REGION Network 8: END: Update the ENO Output. (DO NOT REMOVE. Must be last rung)
   RUNG wire#powerrail
      ReturnCoil( TRUE )
   END_RUNG
   // the same network as SCL:
   ENO := TRUE;
   RETURN;
END_REGION
END_FUNCTION_BLOCK

FUNCTION_BLOCK "UN_07_RecipeControl"   // FB31627, LAD
TITLE = UN_07_RecipeControl
{ S7_Optimized_Access := 'TRUE' }
AUTHOR : tech.team.motioncontrol@siemens.com
FAMILY : CPG
VERSION : 1.0
// Support: tech.team.motioncontrol@siemens.com
   VAR
      instRecipeControl : "CPG_RecipeControl";
      instRecipeManager : "CPG_RecipeHMIManager";
      ONS_RecipeChange : Bool;
      ONS_SaveAsChange : Bool;
      ONS_DeleteChange : Bool;
      ONS_CopyChange : Bool;
   END_VAR
   VAR_TEMP
      tempEnablechange : Bool;
      tempRecipenewname : String[60];
      tempErrorID : Word;
      tempError : Word;
      tempSeconds : Time;
   END_VAR
   VAR CONSTANT
      ERR_CHANGE : Word := 16#8001;
      ERR_SAVE : Word := 16#8002;
      ERR_COPY : Word := 16#8004;
      ERR_DELETE : Word := 16#8008;
   END_VAR
   VAR_TEMP   // added for the SCL form of the ladder/FBD networks
      _w1 : Bool;
      _w2 : Bool;
   END_VAR
BEGIN

REGION Network 1: Determine if recipe change is permitted based on machine state
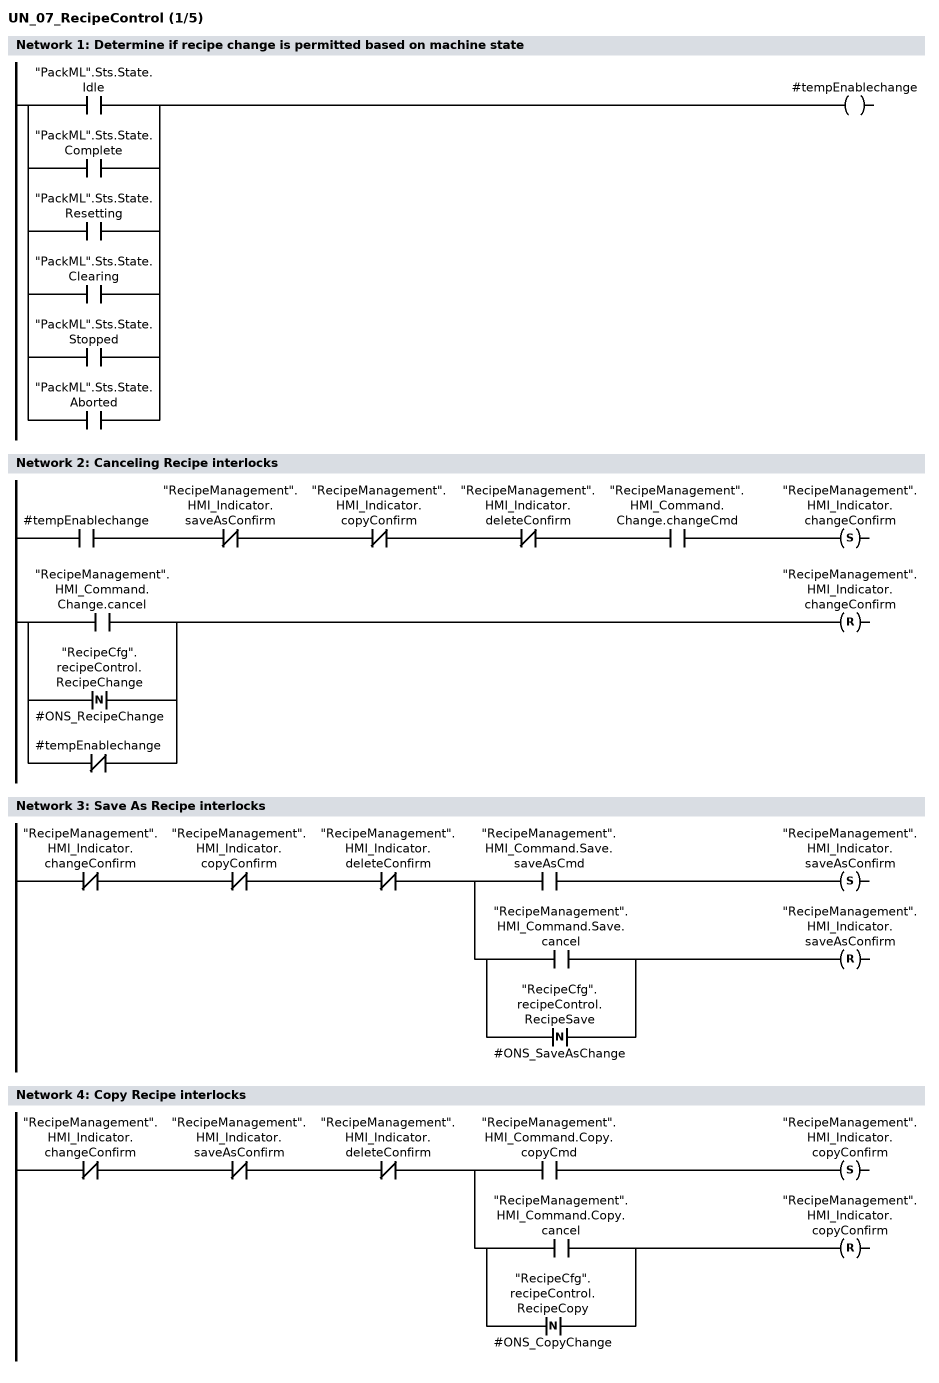
   RUNG wire#powerrail
      Contact( "PackML".Sts.State.Idle )
      wire#w1
      Coil( #tempEnablechange )
   END_RUNG
   RUNG wire#powerrail
      Contact( "PackML".Sts.State.Complete )
   END_RUNG wire#w1
   RUNG wire#powerrail
      Contact( "PackML".Sts.State.Resetting )
   END_RUNG wire#w1
   RUNG wire#powerrail
      Contact( "PackML".Sts.State.Clearing )
   END_RUNG wire#w1
   RUNG wire#powerrail
      Contact( "PackML".Sts.State.Stopped )
   END_RUNG wire#w1
   RUNG wire#powerrail
      Contact( "PackML".Sts.State.Aborted )
   END_RUNG wire#w1
   // the same network as SCL:
   #tempEnablechange := "PackML".Sts.State.Idle OR "PackML".Sts.State.Complete OR "PackML".Sts.State.Resetting OR "PackML".Sts.State.Clearing OR "PackML".Sts.State.Stopped OR "PackML".Sts.State.Aborted;
END_REGION

REGION Network 2: Canceling Recipe interlocks
   RUNG wire#powerrail
      Contact( #tempEnablechange )
      I_Contact( "RecipeManagement".HMI_Indicator.saveAsConfirm )
      I_Contact( "RecipeManagement".HMI_Indicator.copyConfirm )
      I_Contact( "RecipeManagement".HMI_Indicator.deleteConfirm )
      Contact( "RecipeManagement".HMI_Command.Change.changeCmd )
      S_Coil( "RecipeManagement".HMI_Indicator.changeConfirm )
   END_RUNG
   RUNG wire#powerrail
      Contact( "RecipeManagement".HMI_Command.Change.cancel )
      wire#w1
      R_Coil( "RecipeManagement".HMI_Indicator.changeConfirm )
   END_RUNG
   RUNG wire#powerrail
      N_Contact(operand := "RecipeCfg".recipeControl.RecipeChange, bit := #ONS_RecipeChange)
   END_RUNG wire#w1
   RUNG wire#powerrail
      I_Contact( #tempEnablechange )
   END_RUNG wire#w1
   // the same network as SCL:
   IF #tempEnablechange AND NOT "RecipeManagement".HMI_Indicator.saveAsConfirm AND NOT "RecipeManagement".HMI_Indicator.copyConfirm AND NOT "RecipeManagement".HMI_Indicator.deleteConfirm AND "RecipeManagement".HMI_Command.Change.changeCmd THEN
       "RecipeManagement".HMI_Indicator.changeConfirm := TRUE;
   END_IF;
   #_w1 := NOT "RecipeCfg".recipeControl.RecipeChange AND #ONS_RecipeChange;   // falling edge of "RecipeCfg".recipeControl.RecipeChange
   #ONS_RecipeChange := "RecipeCfg".recipeControl.RecipeChange;
   IF "RecipeManagement".HMI_Command.Change.cancel OR #_w1 OR NOT #tempEnablechange THEN
       "RecipeManagement".HMI_Indicator.changeConfirm := FALSE;
   END_IF;
END_REGION

REGION Network 3: Save As Recipe interlocks
   RUNG wire#powerrail
      I_Contact( "RecipeManagement".HMI_Indicator.changeConfirm )
      I_Contact( "RecipeManagement".HMI_Indicator.copyConfirm )
      I_Contact( "RecipeManagement".HMI_Indicator.deleteConfirm )
      wire#w1
      Contact( "RecipeManagement".HMI_Command.Save.saveAsCmd )
      S_Coil( "RecipeManagement".HMI_Indicator.saveAsConfirm )
   END_RUNG
   RUNG wire#w1
      Contact( "RecipeManagement".HMI_Command.Save.cancel )
      wire#w2
      R_Coil( "RecipeManagement".HMI_Indicator.saveAsConfirm )
   END_RUNG
   RUNG wire#w1
      N_Contact(operand := "RecipeCfg".recipeControl.RecipeSave, bit := #ONS_SaveAsChange)
   END_RUNG wire#w2
   // the same network as SCL:
   #_w1 := NOT "RecipeManagement".HMI_Indicator.changeConfirm AND NOT "RecipeManagement".HMI_Indicator.copyConfirm AND NOT "RecipeManagement".HMI_Indicator.deleteConfirm;
   IF #_w1 AND "RecipeManagement".HMI_Command.Save.saveAsCmd THEN
       "RecipeManagement".HMI_Indicator.saveAsConfirm := TRUE;
   END_IF;
   #_w2 := #_w1 AND NOT "RecipeCfg".recipeControl.RecipeSave AND #ONS_SaveAsChange;   // falling edge of "RecipeCfg".recipeControl.RecipeSave
   #ONS_SaveAsChange := "RecipeCfg".recipeControl.RecipeSave;
   IF (#_w1 AND "RecipeManagement".HMI_Command.Save.cancel) OR #_w2 THEN
       "RecipeManagement".HMI_Indicator.saveAsConfirm := FALSE;
   END_IF;
END_REGION

REGION Network 4: Copy Recipe interlocks
   RUNG wire#powerrail
      I_Contact( "RecipeManagement".HMI_Indicator.changeConfirm )
      I_Contact( "RecipeManagement".HMI_Indicator.saveAsConfirm )
      I_Contact( "RecipeManagement".HMI_Indicator.deleteConfirm )
      wire#w1
      Contact( "RecipeManagement".HMI_Command.Copy.copyCmd )
      S_Coil( "RecipeManagement".HMI_Indicator.copyConfirm )
   END_RUNG
   RUNG wire#w1
      Contact( "RecipeManagement".HMI_Command.Copy.cancel )
      wire#w2
      R_Coil( "RecipeManagement".HMI_Indicator.copyConfirm )
   END_RUNG
   RUNG wire#w1
      N_Contact(operand := "RecipeCfg".recipeControl.RecipeCopy, bit := #ONS_CopyChange)
   END_RUNG wire#w2
   // the same network as SCL:
   #_w1 := NOT "RecipeManagement".HMI_Indicator.changeConfirm AND NOT "RecipeManagement".HMI_Indicator.saveAsConfirm AND NOT "RecipeManagement".HMI_Indicator.deleteConfirm;
   IF #_w1 AND "RecipeManagement".HMI_Command.Copy.copyCmd THEN
       "RecipeManagement".HMI_Indicator.copyConfirm := TRUE;
   END_IF;
   #_w2 := #_w1 AND NOT "RecipeCfg".recipeControl.RecipeCopy AND #ONS_CopyChange;   // falling edge of "RecipeCfg".recipeControl.RecipeCopy
   #ONS_CopyChange := "RecipeCfg".recipeControl.RecipeCopy;
   IF (#_w1 AND "RecipeManagement".HMI_Command.Copy.cancel) OR #_w2 THEN
       "RecipeManagement".HMI_Indicator.copyConfirm := FALSE;
   END_IF;
END_REGION

REGION Network 5: Delete Recipe interlocks
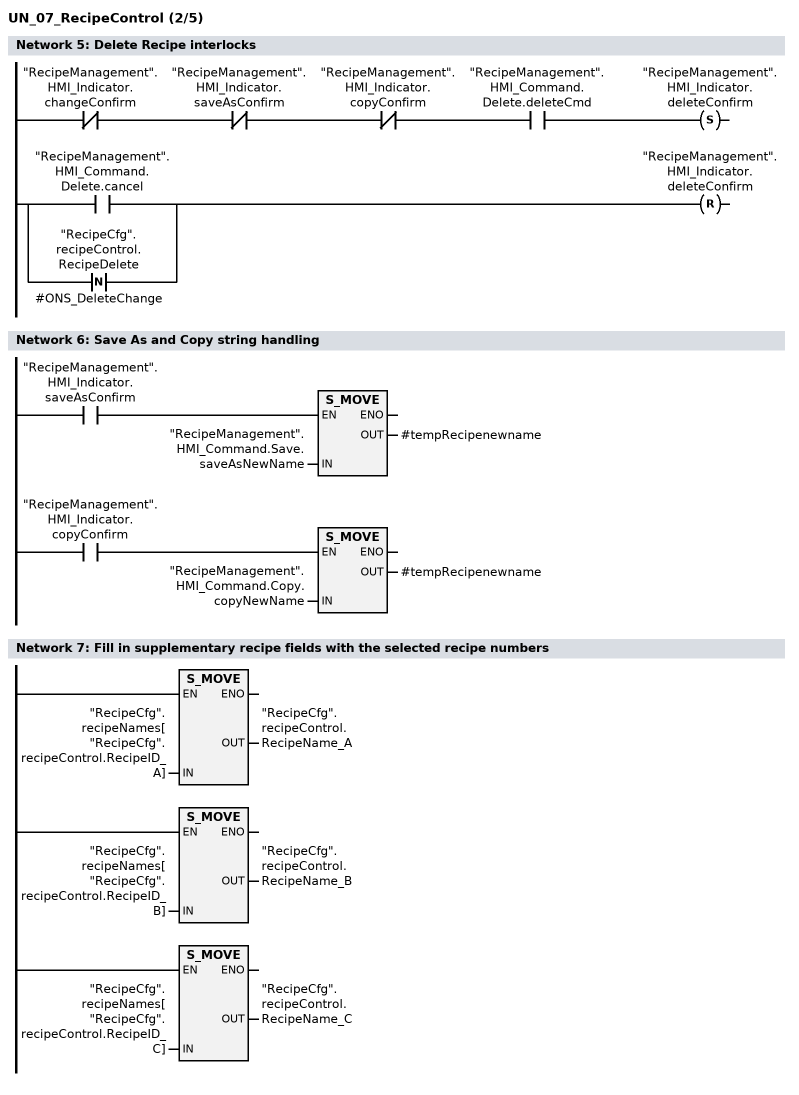
   RUNG wire#powerrail
      I_Contact( "RecipeManagement".HMI_Indicator.changeConfirm )
      I_Contact( "RecipeManagement".HMI_Indicator.saveAsConfirm )
      I_Contact( "RecipeManagement".HMI_Indicator.copyConfirm )
      Contact( "RecipeManagement".HMI_Command.Delete.deleteCmd )
      S_Coil( "RecipeManagement".HMI_Indicator.deleteConfirm )
   END_RUNG
   RUNG wire#powerrail
      Contact( "RecipeManagement".HMI_Command.Delete.cancel )
      wire#w1
      R_Coil( "RecipeManagement".HMI_Indicator.deleteConfirm )
   END_RUNG
   RUNG wire#powerrail
      N_Contact(operand := "RecipeCfg".recipeControl.RecipeDelete, bit := #ONS_DeleteChange)
   END_RUNG wire#w1
   // the same network as SCL:
   IF NOT "RecipeManagement".HMI_Indicator.changeConfirm AND NOT "RecipeManagement".HMI_Indicator.saveAsConfirm AND NOT "RecipeManagement".HMI_Indicator.copyConfirm AND "RecipeManagement".HMI_Command.Delete.deleteCmd THEN
       "RecipeManagement".HMI_Indicator.deleteConfirm := TRUE;
   END_IF;
   #_w1 := NOT "RecipeCfg".recipeControl.RecipeDelete AND #ONS_DeleteChange;   // falling edge of "RecipeCfg".recipeControl.RecipeDelete
   #ONS_DeleteChange := "RecipeCfg".recipeControl.RecipeDelete;
   IF "RecipeManagement".HMI_Command.Delete.cancel OR #_w1 THEN
       "RecipeManagement".HMI_Indicator.deleteConfirm := FALSE;
   END_IF;
END_REGION

REGION Network 6: Save As and Copy string handling
   RUNG wire#powerrail
      Contact( "RecipeManagement".HMI_Indicator.saveAsConfirm )
      S_Move(in := "RecipeManagement".HMI_Command.Save.saveAsNewName, out => #tempRecipenewname)
   END_RUNG
   RUNG wire#powerrail
      Contact( "RecipeManagement".HMI_Indicator.copyConfirm )
      S_Move(in := "RecipeManagement".HMI_Command.Copy.copyNewName, out => #tempRecipenewname)
   END_RUNG
   // the same network as SCL:
   IF "RecipeManagement".HMI_Indicator.saveAsConfirm THEN
       #tempRecipenewname := "RecipeManagement".HMI_Command.Save.saveAsNewName;
   END_IF;
   IF "RecipeManagement".HMI_Indicator.copyConfirm THEN
       #tempRecipenewname := "RecipeManagement".HMI_Command.Copy.copyNewName;
   END_IF;
END_REGION

REGION Network 7: Fill in supplementary recipe fields with the selected recipe numbers
   RUNG wire#powerrail
      S_Move(in := "RecipeCfg".recipeNames["RecipeCfg".recipeControl.RecipeID_A], out => "RecipeCfg".recipeControl.RecipeName_A)
   END_RUNG
   RUNG wire#powerrail
      S_Move(in := "RecipeCfg".recipeNames["RecipeCfg".recipeControl.RecipeID_B], out => "RecipeCfg".recipeControl.RecipeName_B)
   END_RUNG
   RUNG wire#powerrail
      S_Move(in := "RecipeCfg".recipeNames["RecipeCfg".recipeControl.RecipeID_C], out => "RecipeCfg".recipeControl.RecipeName_C)
   END_RUNG
   // the same network as SCL:
   "RecipeCfg".recipeControl.RecipeName_A := "RecipeCfg".recipeNames["RecipeCfg".recipeControl.RecipeID_A];
   "RecipeCfg".recipeControl.RecipeName_B := "RecipeCfg".recipeNames["RecipeCfg".recipeControl.RecipeID_B];
   "RecipeCfg".recipeControl.RecipeName_C := "RecipeCfg".recipeNames["RecipeCfg".recipeControl.RecipeID_C];
END_REGION

REGION Network 8: Call Recipe Control
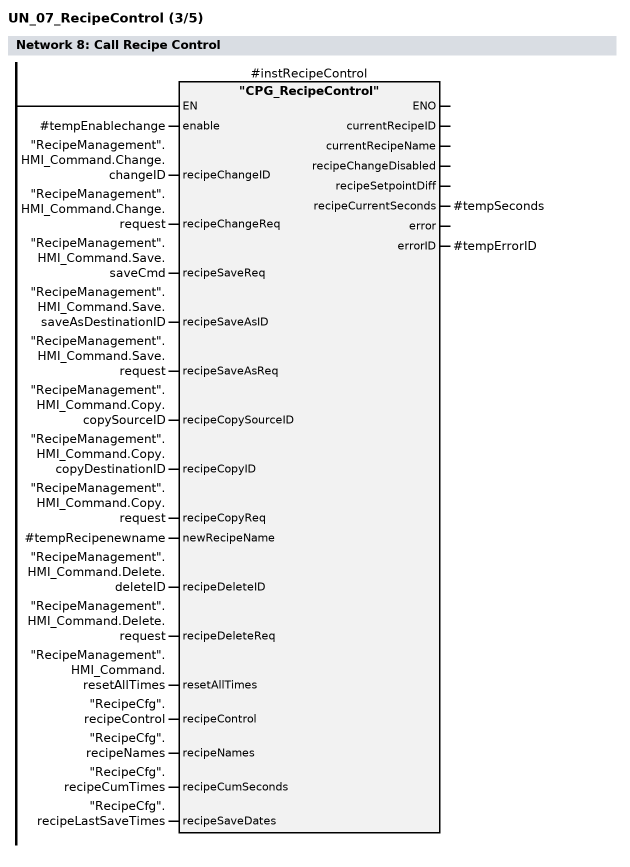
   RUNG wire#powerrail
      #instRecipeControl(enable := #tempEnablechange, recipeChangeID := "RecipeManagement".HMI_Command.Change.changeID, recipeChangeReq := "RecipeManagement".HMI_Command.Change.request, recipeSaveReq := "RecipeManagement".HMI_Command.Save.saveCmd, recipeSaveAsID := "RecipeManagement".HMI_Command.Save.saveAsDestinationID, recipeSaveAsReq := "RecipeManagement".HMI_Command.Save.request, recipeCopySourceID := "RecipeManagement".HMI_Command.Copy.copySourceID, recipeCopyID := "RecipeManagement".HMI_Command.Copy.copyDestinationID, recipeCopyReq := "RecipeManagement".HMI_Command.Copy.request, newRecipeName := #tempRecipenewname, recipeDeleteID := "RecipeManagement".HMI_Command.Delete.deleteID, recipeDeleteReq := "RecipeManagement".HMI_Command.Delete.request, resetAllTimes := "RecipeManagement".HMI_Command.resetAllTimes, recipeControl := "RecipeCfg".recipeControl, recipeNames := "RecipeCfg".recipeNames, recipeCumSeconds := "RecipeCfg".recipeCumTimes, recipeSaveDates := "RecipeCfg".recipeLastSaveTimes, currentRecipeID =>, currentRecipeName =>, recipeChangeDisabled =>, recipeSetpointDiff =>, recipeCurrentSeconds => #tempSeconds, error =>, errorID => #tempErrorID)
   END_RUNG
   // the same network as SCL:
   #instRecipeControl(enable := #tempEnablechange,   // "CPG_RecipeControl"
                      recipeChangeID := "RecipeManagement".HMI_Command.Change.changeID,
                      recipeChangeReq := "RecipeManagement".HMI_Command.Change.request,
                      recipeSaveReq := "RecipeManagement".HMI_Command.Save.saveCmd,
                      recipeSaveAsID := "RecipeManagement".HMI_Command.Save.saveAsDestinationID,
                      recipeSaveAsReq := "RecipeManagement".HMI_Command.Save.request,
                      recipeCopySourceID := "RecipeManagement".HMI_Command.Copy.copySourceID,
                      recipeCopyID := "RecipeManagement".HMI_Command.Copy.copyDestinationID,
                      recipeCopyReq := "RecipeManagement".HMI_Command.Copy.request,
                      newRecipeName := #tempRecipenewname,
                      recipeDeleteID := "RecipeManagement".HMI_Command.Delete.deleteID,
                      recipeDeleteReq := "RecipeManagement".HMI_Command.Delete.request,
                      resetAllTimes := "RecipeManagement".HMI_Command.resetAllTimes,
                      recipeControl := "RecipeCfg".recipeControl,
                      recipeNames := "RecipeCfg".recipeNames,
                      recipeCumSeconds := "RecipeCfg".recipeCumTimes,
                      recipeSaveDates := "RecipeCfg".recipeLastSaveTimes,
                      recipeCurrentSeconds => #tempSeconds,
                      errorID => #tempErrorID);
END_REGION

REGION Network 9: Clear IDs from HMI if not on that screen
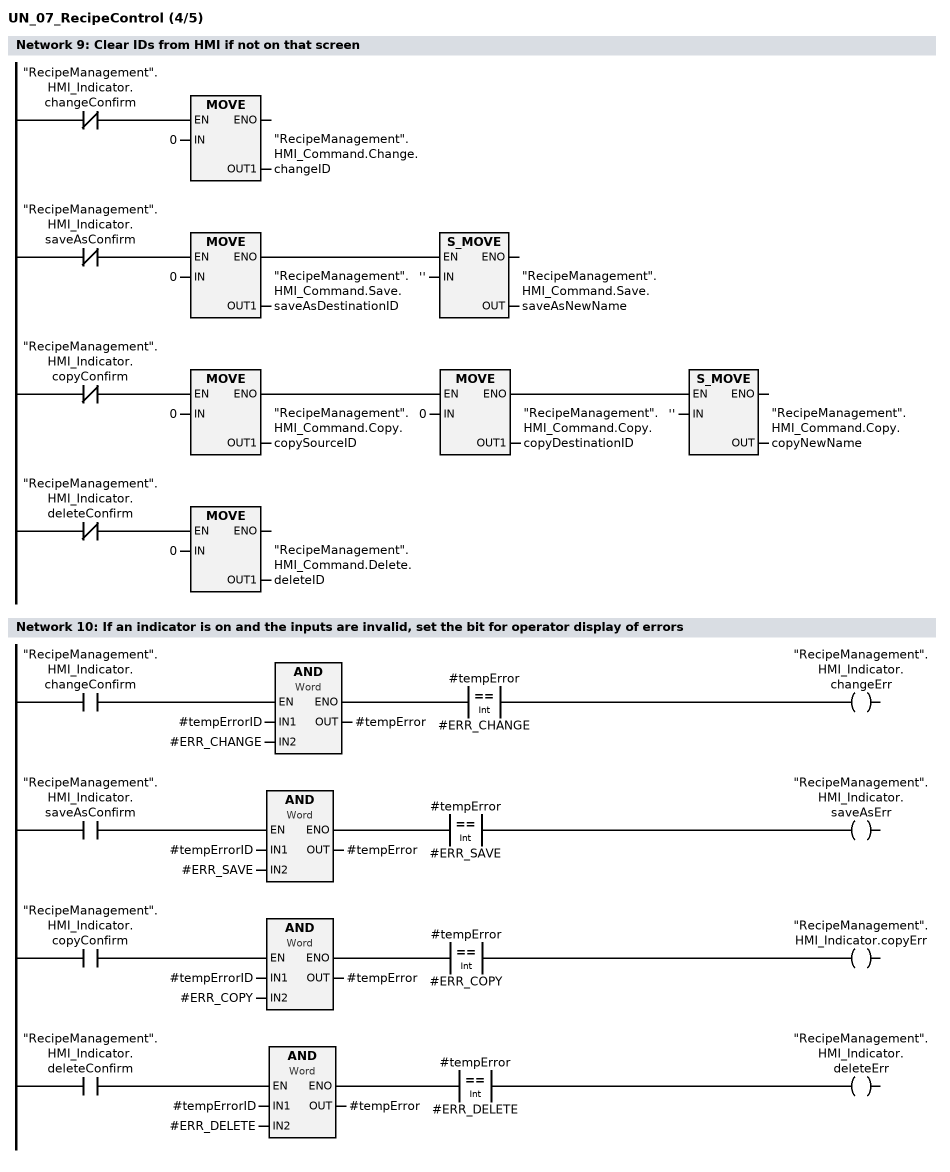
   RUNG wire#powerrail
      I_Contact( "RecipeManagement".HMI_Indicator.changeConfirm )
      Move(in := 0, out1 => "RecipeManagement".HMI_Command.Change.changeID)
   END_RUNG
   RUNG wire#powerrail
      I_Contact( "RecipeManagement".HMI_Indicator.saveAsConfirm )
      Move(in := 0, out1 => "RecipeManagement".HMI_Command.Save.saveAsDestinationID)
      S_Move(in := '', out => "RecipeManagement".HMI_Command.Save.saveAsNewName)
   END_RUNG
   RUNG wire#powerrail
      I_Contact( "RecipeManagement".HMI_Indicator.copyConfirm )
      Move(in := 0, out1 => "RecipeManagement".HMI_Command.Copy.copySourceID)
      Move(in := 0, out1 => "RecipeManagement".HMI_Command.Copy.copyDestinationID)
      S_Move(in := '', out => "RecipeManagement".HMI_Command.Copy.copyNewName)
   END_RUNG
   RUNG wire#powerrail
      I_Contact( "RecipeManagement".HMI_Indicator.deleteConfirm )
      Move(in := 0, out1 => "RecipeManagement".HMI_Command.Delete.deleteID)
   END_RUNG
   // the same network as SCL:
   IF NOT "RecipeManagement".HMI_Indicator.changeConfirm THEN
       "RecipeManagement".HMI_Command.Change.changeID := 0;
   END_IF;
   IF NOT "RecipeManagement".HMI_Indicator.saveAsConfirm THEN
       "RecipeManagement".HMI_Command.Save.saveAsDestinationID := 0;
       "RecipeManagement".HMI_Command.Save.saveAsNewName := '';
   END_IF;
   IF NOT "RecipeManagement".HMI_Indicator.copyConfirm THEN
       "RecipeManagement".HMI_Command.Copy.copySourceID := 0;
       "RecipeManagement".HMI_Command.Copy.copyDestinationID := 0;
       "RecipeManagement".HMI_Command.Copy.copyNewName := '';
   END_IF;
   IF NOT "RecipeManagement".HMI_Indicator.deleteConfirm THEN
       "RecipeManagement".HMI_Command.Delete.deleteID := 0;
   END_IF;
END_REGION

REGION Network 10: If an indicator is on and the inputs are invalid, set the bit for operator display of errors
   RUNG wire#powerrail
      Contact( "RecipeManagement".HMI_Indicator.changeConfirm )
      { S7_Templates := "SrcType := Word" } And(in1 := #tempErrorID, in2 := #ERR_CHANGE, out => #tempError)
      { S7_Templates := "SrcType := Int" } EQ_Contact(in1 := #tempError, in2 := #ERR_CHANGE)
      Coil( "RecipeManagement".HMI_Indicator.changeErr )
   END_RUNG
   RUNG wire#powerrail
      Contact( "RecipeManagement".HMI_Indicator.saveAsConfirm )
      { S7_Templates := "SrcType := Word" } And(in1 := #tempErrorID, in2 := #ERR_SAVE, out => #tempError)
      { S7_Templates := "SrcType := Int" } EQ_Contact(in1 := #tempError, in2 := #ERR_SAVE)
      Coil( "RecipeManagement".HMI_Indicator.saveAsErr )
   END_RUNG
   RUNG wire#powerrail
      Contact( "RecipeManagement".HMI_Indicator.copyConfirm )
      { S7_Templates := "SrcType := Word" } And(in1 := #tempErrorID, in2 := #ERR_COPY, out => #tempError)
      { S7_Templates := "SrcType := Int" } EQ_Contact(in1 := #tempError, in2 := #ERR_COPY)
      Coil( "RecipeManagement".HMI_Indicator.copyErr )
   END_RUNG
   RUNG wire#powerrail
      Contact( "RecipeManagement".HMI_Indicator.deleteConfirm )
      { S7_Templates := "SrcType := Word" } And(in1 := #tempErrorID, in2 := #ERR_DELETE, out => #tempError)
      { S7_Templates := "SrcType := Int" } EQ_Contact(in1 := #tempError, in2 := #ERR_DELETE)
      Coil( "RecipeManagement".HMI_Indicator.deleteErr )
   END_RUNG
   // the same network as SCL:
   IF "RecipeManagement".HMI_Indicator.changeConfirm THEN #tempError := #tempErrorID AND #ERR_CHANGE; END_IF;
   "RecipeManagement".HMI_Indicator.changeErr := "RecipeManagement".HMI_Indicator.changeConfirm AND (#tempError = #ERR_CHANGE);
   IF "RecipeManagement".HMI_Indicator.saveAsConfirm THEN #tempError := #tempErrorID AND #ERR_SAVE; END_IF;
   "RecipeManagement".HMI_Indicator.saveAsErr := "RecipeManagement".HMI_Indicator.saveAsConfirm AND (#tempError = #ERR_SAVE);
   IF "RecipeManagement".HMI_Indicator.copyConfirm THEN #tempError := #tempErrorID AND #ERR_COPY; END_IF;
   "RecipeManagement".HMI_Indicator.copyErr := "RecipeManagement".HMI_Indicator.copyConfirm AND (#tempError = #ERR_COPY);
   IF "RecipeManagement".HMI_Indicator.deleteConfirm THEN #tempError := #tempErrorID AND #ERR_DELETE; END_IF;
   "RecipeManagement".HMI_Indicator.deleteErr := "RecipeManagement".HMI_Indicator.deleteConfirm AND (#tempError = #ERR_DELETE);
END_REGION

REGION Network 11: Call Recipe HMI Manager to handle display of setpoints
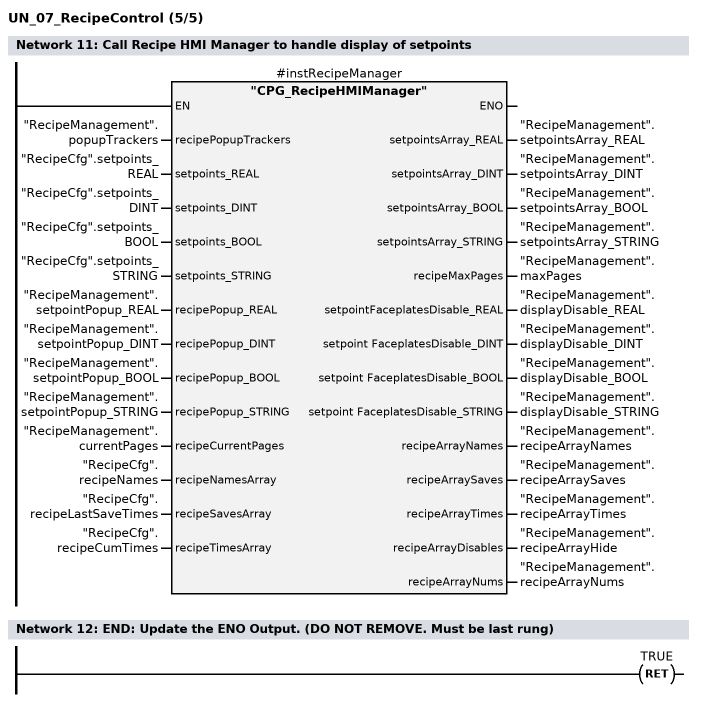
   RUNG wire#powerrail
      #instRecipeManager(recipePopupTrackers := "RecipeManagement".popupTrackers, setpoints_REAL := "RecipeCfg".setpoints_REAL, setpoints_DINT := "RecipeCfg".setpoints_DINT, setpoints_BOOL := "RecipeCfg".setpoints_BOOL, setpoints_STRING := "RecipeCfg".setpoints_STRING, recipePopup_REAL := "RecipeManagement".setpointPopup_REAL, recipePopup_DINT := "RecipeManagement".setpointPopup_DINT, recipePopup_BOOL := "RecipeManagement".setpointPopup_BOOL, recipePopup_STRING := "RecipeManagement".setpointPopup_STRING, recipeCurrentPages := "RecipeManagement".currentPages, recipeNamesArray := "RecipeCfg".recipeNames, recipeSavesArray := "RecipeCfg".recipeLastSaveTimes, recipeTimesArray := "RecipeCfg".recipeCumTimes, setpointsArray_REAL => "RecipeManagement".setpointsArray_REAL, setpointsArray_DINT => "RecipeManagement".setpointsArray_DINT, setpointsArray_BOOL => "RecipeManagement".setpointsArray_BOOL, setpointsArray_STRING => "RecipeManagement".setpointsArray_STRING, recipeMaxPages => "RecipeManagement".maxPages, setpointFaceplatesDisable_REAL => "RecipeManagement".displayDisable_REAL, "setpoint FaceplatesDisable_DINT" => "RecipeManagement".displayDisable_DINT, "setpoint FaceplatesDisable_BOOL" => "RecipeManagement".displayDisable_BOOL, "setpoint FaceplatesDisable_STRING" => "RecipeManagement".displayDisable_STRING, recipeArrayNames => "RecipeManagement".recipeArrayNames, recipeArraySaves => "RecipeManagement".recipeArraySaves, recipeArrayTimes => "RecipeManagement".recipeArrayTimes, recipeArrayDisables => "RecipeManagement".recipeArrayHide, recipeArrayNums => "RecipeManagement".recipeArrayNums)
   END_RUNG
   // the same network as SCL:
   #instRecipeManager(recipePopupTrackers := "RecipeManagement".popupTrackers,   // "CPG_RecipeHMIManager"
                      setpoints_REAL := "RecipeCfg".setpoints_REAL,
                      setpoints_DINT := "RecipeCfg".setpoints_DINT,
                      setpoints_BOOL := "RecipeCfg".setpoints_BOOL,
                      setpoints_STRING := "RecipeCfg".setpoints_STRING,
                      recipePopup_REAL := "RecipeManagement".setpointPopup_REAL,
                      recipePopup_DINT := "RecipeManagement".setpointPopup_DINT,
                      recipePopup_BOOL := "RecipeManagement".setpointPopup_BOOL,
                      recipePopup_STRING := "RecipeManagement".setpointPopup_STRING,
                      recipeCurrentPages := "RecipeManagement".currentPages,
                      recipeNamesArray := "RecipeCfg".recipeNames,
                      recipeSavesArray := "RecipeCfg".recipeLastSaveTimes,
                      recipeTimesArray := "RecipeCfg".recipeCumTimes,
                      setpointsArray_REAL => "RecipeManagement".setpointsArray_REAL,
                      setpointsArray_DINT => "RecipeManagement".setpointsArray_DINT,
                      setpointsArray_BOOL => "RecipeManagement".setpointsArray_BOOL,
                      setpointsArray_STRING => "RecipeManagement".setpointsArray_STRING,
                      recipeMaxPages => "RecipeManagement".maxPages,
                      setpointFaceplatesDisable_REAL => "RecipeManagement".displayDisable_REAL,
                      "setpoint FaceplatesDisable_DINT" => "RecipeManagement".displayDisable_DINT,
                      "setpoint FaceplatesDisable_BOOL" => "RecipeManagement".displayDisable_BOOL,
                      "setpoint FaceplatesDisable_STRING" => "RecipeManagement".displayDisable_STRING,
                      recipeArrayNames => "RecipeManagement".recipeArrayNames,
                      recipeArraySaves => "RecipeManagement".recipeArraySaves,
                      recipeArrayTimes => "RecipeManagement".recipeArrayTimes,
                      recipeArrayDisables => "RecipeManagement".recipeArrayHide,
                      recipeArrayNums => "RecipeManagement".recipeArrayNums);
END_REGION

REGION Network 12: END: Update the ENO Output. (DO NOT REMOVE. Must be last rung)
   RUNG wire#powerrail
      ReturnCoil( TRUE )
   END_RUNG
   // the same network as SCL:
   ENO := TRUE;
   RETURN;
END_REGION
END_FUNCTION_BLOCK

// ===== library types =====

// folder: ISA_TR88/CPG_Types

TYPE "UDT_TR88_CPG_EventStatus"
AUTHOR : FoodBev
FAMILY : ISATR88e
NAME : EventSts
VERSION : 1.0
   STRUCT
      Sts_FirstOutEvent : "UDT_TR88_CPG_Event";   // Event Info of the very first active event (irregardeless of the cat)
      Sts_FirstOutEventCat : Array[0..9] of "UDT_TR88_CPG_Event";
      Sts_Events : Array[0.."TR88_CPG_NoOfStsElements_EventStatus"] of "UDT_TR88_CPG_Event";
      Sts_NumEvents : Int;   // number of all current active events
      Sts_NumAllEvents : Int;   // number of all current events
      Out_ZeroEvent : "UDT_TR88_CPG_Event";   // null event information
      Sts_Category_0_Latched : Bool;   // Category 0 Event - latched (require reset cmd)
      Sts_Category_1_Latched : Bool;   // Category 1 Event - latched (require reset cmd)
      Sts_Category_2_Latched : Bool;   // Category 2 Event - latched (require reset cmd)
      Sts_Category_3_Latched : Bool;   // Category 3 Event - latched (require reset cmd)
      Sts_Category_4_Latched : Bool;   // Category 4 Event - latched (require reset cmd)
      Sts_Category_5_Latched : Bool;   // Category 5 Event - latched (require reset cmd)
      Sts_Category_6_Latched : Bool;   // Category 6 Event - latched (require reset cmd)
      Sts_Category_7_Latched : Bool;   // Category 7 Event - latched (require reset cmd)
      Sts_Category_8_Latched : Bool;   // Category 8 Event - latched (require reset cmd)
      Sts_Category_9_Latched : Bool;   // Category 9 Event - latched (require reset cmd)
      Sts_Category_0_NotLatched : Bool;   // Category 0 Event - NotLatched (currently active)
      Sts_Category_1_NotLatched : Bool;   // Category 1 Event - NotLatched (currently active)
      Sts_Category_2_NotLatched : Bool;   // Category 2 Event - NotLatched (currently active)
      Sts_Category_3_NotLatched : Bool;   // Category 3 Event - NotLatched (currently active)
      Sts_Category_4_NotLatched : Bool;   // Category 4 Event - NotLatched (currently active)
      Sts_Category_5_NotLatched : Bool;   // Category 5 Event - NotLatched (currently active)
      Sts_Category_6_NotLatched : Bool;   // Category 6 Event - NotLatched (currently active)
      Sts_Category_7_NotLatched : Bool;   // Category 7 Event - NotLatched (currently active)
      Sts_Category_8_NotLatched : Bool;   // Category 8 Event - NotLatched (currently active)
      Sts_Category_9_NotLatched : Bool;   // Category 9 Event - NotLatched (currently active)
      Sts_CurrentActiveEvent : Bool;   // Active # of Event
      Wrk_ResetID : Int;   // Working Variable - DO NOT MODIFY
      Wrk_EventArraySize : Int;   // Working Variable - DO NOT MODIFY
      Wrk_UpdateEventListID : Int;   // Working Variable - DO NOT MODIFY
      Wrk_LanguageSelection : Int;   // This is the value of language selected in the HMI
      Wrk_MessagePrefix : String[10];   // Working Variable - DO NOT MODIFY
   END_STRUCT;
END_TYPE

TYPE "UDT_TR88_CPG_EventCfg"
AUTHOR : FoodBev
FAMILY : ISATR88e
NAME : EvntCfgA
VERSION : 1.0
   STRUCT
      ID : Int;   // ID Value - from PackTags Reason Code, 1=E-Stop pushed, 3=Main off, etc.
      Value : Int;   // Reason Code 'Value' - allows for detailed breakdown of ID, ie 1=Discharge,
      Message : Array[0.."LPMLV30_LANGUAGES_UPPER_LIM"] of String["TR88_CPG_MsgEventStringLength"];   // Alarm Message - 0=English,1=Spanish, 2=German, 3=Italian, 4=French
      Category : Int;   // Category Value (0-9)
   END_STRUCT;
END_TYPE

TYPE "UDT_TR88_CPG_Event"
AUTHOR : FoodBev
FAMILY : ISATR88e
NAME : Event
VERSION : 1.0
   STRUCT
      Trigger : Bool;   // Internal trigger bit
      ID : Int;   // ID Value - from PackTags Reason Code, 1=E-Stop pushed, 3=Main off, etc
      Value : Int;   // Reason Code 'Value' - allows for detailed breakdown of ID, ie 1=Discharge
      Message : String["TR88_CPG_MsgEventStringLength"];   // Message OF alarm = prefix message + alarm message
      Category : Int;   // Category Value (0-9)
      DateTime : DTL;   // Time & date (DTL) the event was initially triggered
      AckDateTime : DTL;   // Time & date (DTL) the event was acknowledged
   END_STRUCT;
END_TYPE

TYPE "UDT_TR88_CPG_EventSummation"
AUTHOR : FoodBev
FAMILY : ISATR88e
NAME : EventSum
VERSION : 1.0
   STRUCT
      Sts_FirstOutEvent : "UDT_TR88_CPG_Event";   // First Out (Stop Reason) Event
      Sts_FirstOutEventCat : Array[0..9] of "UDT_TR88_CPG_Event";   // First Out (Stop Reason) Event by Category\
      Sts_Events : Array[0.."TR88_CPG_NoOfStsElements_EventSum"] of "UDT_TR88_CPG_Event";   // All Active Events
      Sts_NumEvents : Int;   // Number of Active Events
      Sts_Category_0_Latched : Bool;   // Category 0 Event - latched (require reset cmd)
      Sts_Category_1_Latched : Bool;   // Category 1 Event - latched (require reset cmd)
      Sts_Category_2_Latched : Bool;   // Category 2 Event - latched (require reset cmd)
      Sts_Category_3_Latched : Bool;   // Category 3 Event - latched (require reset cmd)
      Sts_Category_4_Latched : Bool;   // Category 4 Event - latched (require reset cmd)
      Sts_Category_5_Latched : Bool;   // Category 5 Event - latched (require reset cmd)
      Sts_Category_6_Latched : Bool;   // Category 6 Event - latched (require reset cmd)
      Sts_Category_7_Latched : Bool;   // Category 7 Event - latched (require reset cmd)
      Sts_Category_8_Latched : Bool;   // Category 8 Event - latched (require reset cmd)
      Sts_Category_9_Latched : Bool;   // Category 9 Event - latched (require reset cmd)
      Sts_Category_0_NotLatched : Bool;   // Category 0 Event - NotLatched (currently active)
      Sts_Category_1_NotLatched : Bool;   // Category 1 Event - NotLatched (currently active)
      Sts_Category_2_NotLatched : Bool;   // Category 2 Event - NotLatched (currently active)
      Sts_Category_3_NotLatched : Bool;   // Category 3 Event - NotLatched (currently active)
      Sts_Category_4_NotLatched : Bool;   // Category 4 Event - NotLatched (currently active)
      Sts_Category_5_NotLatched : Bool;   // Category 5 Event - NotLatched (currently active)
      Sts_Category_6_NotLatched : Bool;   // Category 6 Event - NotLatched (currently active)
      Sts_Category_7_NotLatched : Bool;   // Category 7 Event - NotLatched (currently active)
      Sts_Category_8_NotLatched : Bool;   // Category 8 Event - NotLatched (currently active)
      Sts_Category_9_NotLatched : Bool;   // Category 9 Event - NotLatched (currently active)
      Sts_CurrentActiveEvent : Bool;   // Event Active = 1, not active = 0
      Wrk_EventArraySize : Int;   // Maximum Array Size - DO NOT MODIFY
      Wrk_Category_0_Latched : Bool;   // Working Variable - DO NOT MODIFY
      Wrk_Category_1_Latched : Bool;   // Working Variable - DO NOT MODIFY
      Wrk_Category_2_Latched : Bool;   // Working Variable - DO NOT MODIFY
      Wrk_Category_3_Latched : Bool;   // Working Variable - DO NOT MODIFY
      Wrk_Category_4_Latched : Bool;   // Working Variable - DO NOT MODIFY
      Wrk_Category_5_Latched : Bool;   // Working Variable - DO NOT MODIFY
      Wrk_Category_6_Latched : Bool;   // Working Variable - DO NOT MODIFY
      Wrk_Category_7_Latched : Bool;   // Working Variable - DO NOT MODIFY
      Wrk_Category_8_Latched : Bool;   // Working Variable - DO NOT MODIFY
      Wrk_Category_9_Latched : Bool;   // Working Variable - DO NOT MODIFY
      Wrk_Category_0_NotLatched : Bool;   // Working Variable - DO NOT MODIFY
      Wrk_Category_1_NotLatched : Bool;   // Working Variable - DO NOT MODIFY
      Wrk_Category_2_NotLatched : Bool;   // Working Variable - DO NOT MODIFY
      Wrk_Category_3_NotLatched : Bool;   // Working Variable - DO NOT MODIFY
      Wrk_Category_4_NotLatched : Bool;   // Working Variable - DO NOT MODIFY
      Wrk_Category_5_NotLatched : Bool;   // Working Variable - DO NOT MODIFY
      Wrk_Category_6_NotLatched : Bool;   // Working Variable - DO NOT MODIFY
      Wrk_Category_7_NotLatched : Bool;   // Working Variable - DO NOT MODIFY
      Wrk_Category_8_NotLatched : Bool;   // Working Variable - DO NOT MODIFY
      Wrk_Category_9_NotLatched : Bool;   // Working Variable - DO NOT MODIFY
      Wrk_CurrentActiveEvent : Bool;   // Working Variable - DO NOT MODIFY
   END_STRUCT;
END_TYPE

TYPE "UDT_TR88_CPG_PackML_Module_Sts"
AUTHOR : FoodBev
FAMILY : ISATR88e
NAME : PML_MdSt
VERSION : 1.0
   STRUCT
      Cmd_Reset : Bool;   // Reset
      Sts_Resetting_SC : Bool;   // Resetting State Complete
      Cmd_Start : Bool;   // Start
      Sts_Starting_SC : Bool;   // Starting State Complete
      Cmd_Stop : Bool;   // Stop
      Sts_Stopping_SC : Bool;   // Stopping State Complete
      Cmd_Hold : Bool;   // Hold
      Sts_Holding_SC : Bool;   // Holding State Complete
      Cmd_UnHold : Bool;   // UnHold
      Sts_UnHolding_SC : Bool;   // UnHolding State Complete
      Cmd_Suspend : Bool;   // Suspend
      Sts_Suspending_SC : Bool;   // Suspending State Complete
      Cmd_UnSuspend : Bool;   // UnSuspend
      Sts_UnSuspending_SC : Bool;   // UnSuspending State Complete
      Cmd_Abort : Bool;   // Abort
      Sts_Aborting_SC : Bool;   // Aborting State Complete
      Cmd_Clear : Bool;   // Clear
      Sts_Clearing_SC : Bool;   // Clearing State Complete
      Sts_Execute_SC : Bool;   // Execute State Complete
      Sts_Completing_SC : Bool;   // Completing State Complete
      ModuleActive : Bool;   // Module Active Bit
      ONS : Bool;   // OneShot bit
   END_STRUCT;
END_TYPE

TYPE "UDT_TR88_CPG_Message_Prefix"
VERSION : 0.1
   STRUCT
      MessagePrefix : Array[0.."LPMLV30_LANGUAGES_UPPER_LIM"] of String["TR88_CPG_MsgPrefixStringLength"];   // Multi-Lingual Messagage for Prefix (i.e 0=EN, 1=SP/ES, 2=DE, 3=FR, 4=IT)
   END_STRUCT;
END_TYPE

TYPE "UDT_TR88_CPG_Message_Event"
VERSION : 0.1
   STRUCT
      Language : Array[0.."LPMLV30_LANGUAGES_UPPER_LIM"] of String["TR88_CPG_MsgEventStringLength"];   // Multi-Lingual Message for Events Msg (i.e 0=EN, 1=SP/ES, 2=DE, 3=FR, 4=IT)
   END_STRUCT;
END_TYPE

// folder: ISA_TR88/CPG_Blocks

FUNCTION_BLOCK "FB_TR88_CPG_Event"   // FB3101, SCL
TITLE = PackML Event (TR88 CPG Template)
{ S7_Optimized_Access := 'TRUE' }
AUTHOR : FoodBev
FAMILY : ISATR88e
NAME : Event
VERSION : 2.0
// This FB, designed to have minimal impact on scan time, resides inside the control module code. Whenever rung conditions preceding this FB are true, then the event configuration is copied to the equipment modules input event list and the event is latched on with the controller time. When the rung conditions are false, the event will stay latched until a reset command is sent. Each instance of this FB corresponds to a different event. For example, if a control module generates 2 faults, then this FB will be programmed twice in the control module routine. Each event can also belong to a category, from 0-9, for grouping or prioritizing event information for reporting purposed.
   VAR_INPUT
      EnableIn : Bool;   // Enable the FB call.
      Cfg_Event : "UDT_TR88_CPG_EventCfg";   // configuration data structure for this event
      Cfg_MessagePrefix : "UDT_TR88_CPG_Message_Prefix";   // Message Prefix value for event messages
   END_VAR
   VAR_OUTPUT
      Sts_Active : Bool;   // event is currently active
      Sts_Latched : Bool;   // event has been active since last reset command
   END_VAR
   VAR_IN_OUT
      In_EventStatus : "UDT_TR88_CPG_EventStatus";   // Working event list data section
   END_VAR
   VAR
      Event_Number : Int;   // Event Number
      Prev_ResetID : Int;   // Prev Reset ID
      error_RTC : Int;   // Error code for reading of Real Time Clock
      Event_CurDateTime : Date_And_Time;   // temp value for current date & time
   END_VAR
   VAR_TEMP
      "step" : Int;
      temp_text1 : String[30];   // temp string value
      temp_text2 : String[30];   // temp string value
      temp_text3 : String[30];   // temp string value
      temp_Language : Int;   // value of the currently selected langauge
   END_VAR
BEGIN
   // ============================================================================ 
   // FUNCTION_BLOCK "FB_PMLe_Event"
   // ---------------------------------------------------------------------------
   // Siemens Industry, Inc.
   // Food & Beverage VSS
   // ---------------------------------------------------------------------------
   // FUNCTIONALITY:  
   // Function Block to control TR88 EVENT functions for CPG Template. 
   // ---------------------------------------------------------------------------
   // change log table:
   // version        date          expert in charge        changes applied
   //  1.6       2012.02.01        Mike Pieper        Inital Release - Rev 1.6 
   //  1.7       2013.07.31        Mike Pieper        Fixed bug for EM message prefix
   //  2.0       2015.04.01        Mike Pieper        TR88.00.02 Edition 2 Release. 
   //  =========================================================================== 
   (*
   THIS SOFTWARE IS PROVIDED "AS IS" AND WITHOUT WARRANTIES OF ANY KIND, WHETHER EXPRESS OR IMPLIED.

   General information -
       Note :  the standard applications are NOT binding AND DO NOT claim TO be complete regarding configuration, equipment OR any eventuality which may arise. 
       The standard applications DO NOT represent specific customer solutions, but are only intended TO provide support FOR typical tasks. You are responsible 
       FOR the proper operation OF the described products. These standard applications DO NOT relieve you OF your responsibility regarding the safe handling 
       when using, installing operating AND maintaining the equipment. BY using these standard applications, you agree that Siemens cannot be made liable FOR 
       possible damage beyond the mentioned liability clause. We reserve the right TO make changes AND revisions TO these standard applications at Any Time 
       without prior notice. In the CASE OF Any differences between the suggestions made in these standard applications AND other publications from Siemens, 
       such as catalogs, the contents OF the other documentation have priority.

   Warranty conditions, liability, AND support -
      IF the application has been made available free OF charge, the following applies:
      * We DO NOT provide a warranty FOR Any OF the information contained in this document.
      * All other rights AND claims against Siemens AG irrespective OF legal basis are excluded. In particular claims FOR damages against Siemens AG 
      in the CASE OF Product outage, downtime, loss OF profit, either directly, indirectly OR consequential damage are excluded.
      * This does NOT apply when liability is compulsory BY law, e. g. in the CASE OF the Product liability act, premeditation, an act OF gross negligence 
      BY superiors AND managerial staff OF Siemens AG OR in cases OF fraudulent concealment OF defects.
      * This limitation OF liability also applies TO sub-contractors, suppliers, delegates, superiors AND managerial staff OF Siemens AG.
      German law shall apply TO this agreement FOR customers with head offices in Germany; Swiss law FOR customers with head offices outside Germany. 
      Application OF the United Nations Convention on Contracts FOR the International Sale OF Goods as OF 11.04.1980 (CISG) is excluded.
   *)

   // ===========================================================================
   //  Begin the LOGIC section:

   //-------------  If ENABLE is FALSE----------------------------------------
   IF NOT(#EnableIn)                          // If block is not enabled, then
       THEN             
           IF #Sts_Active THEN              // Status Active
               IF #Event_Number < #In_EventStatus.Wrk_EventArraySize THEN   // current event below max size?
                   #error_RTC := RD_LOC_T (OUT=> #Event_CurDateTime);            // Read the Real Time Clock with local time settings
                   #In_EventStatus.Sts_Events[#Event_Number].AckDateTime := #Event_CurDateTime; // update Acknowledge time
                   #In_EventStatus.Sts_Events[#Event_Number].Trigger := false;
               END_IF;                     // IF Event_Number

               #Sts_Active:= false;             // Reset the active bit        
               #In_EventStatus.Wrk_UpdateEventListID := #In_EventStatus.Wrk_UpdateEventListID+1;
           END_IF;                             // IF Sts_Active

           IF #Sts_Latched AND (#In_EventStatus.Wrk_ResetID <> #Prev_ResetID) THEN
               #Sts_Latched :=false;
               #In_EventStatus.Wrk_UpdateEventListID := #In_EventStatus.Wrk_UpdateEventListID+1;
               #Prev_ResetID := #In_EventStatus.Wrk_ResetID;
           END_IF;             // IF Sts_Latched

           ENO:= FALSE;         // enable out is false (0)
   ELSE                    // else IF NOT (enable)

   //-------------  If ENABLE is TRUE ----------------------------------------  
   // If this FB is enabled....  
   IF NOT (#Sts_Active) OR (#In_EventStatus.Wrk_ResetID <> #Prev_ResetID) THEN
       IF NOT (#Sts_Latched)  THEN
           #error_RTC := RD_LOC_T (OUT=> #Event_CurDateTime);            // Read the Real Time Clock using local time settings      
       END_IF;

       IF NOT (#Sts_Latched) OR (#In_EventStatus.Wrk_ResetID <> #Prev_ResetID) THEN
           #Event_Number                    := #In_EventStatus.Sts_NumAllEvents;             // increment event number
           #In_EventStatus.Sts_NumAllEvents := #In_EventStatus.Sts_NumAllEvents + 1;         // increment number of all event
           #Prev_ResetID := #In_EventStatus.Wrk_ResetID;                                     // update previous Reset ID      
       END_IF;

      IF #Event_Number < #In_EventStatus.Wrk_EventArraySize THEN    
           #temp_Language := #In_EventStatus.Wrk_LanguageSelection;

           #In_EventStatus.Sts_Events[#Event_Number].ID         := #Cfg_Event.ID;
           #In_EventStatus.Sts_Events[#Event_Number].Value      := #Cfg_Event.Value;
           #In_EventStatus.Sts_Events[#Event_Number].Category   := #Cfg_Event.Category;

           // V2.0 changess
           // = Inp_EventStatus.Sts_Events[#Event_Number].Message := Inp_EventStatus.Wrk_MessagePrefix + #Cfg_MessagePrefix[Inp_EventStatus.Wrk_LanguageSelection]+ #Cfg_Event.Message[Inp_EventStatus.Wrk_LanguageSelection]
           // Ensure sure that strings have a valid character.  If null(zero) length, then CONCAT will generate an error, thus a filler (space or _) prevents this problem
           #temp_text1 := #In_EventStatus.Wrk_MessagePrefix;
           IF LEN(#temp_text1) = 0 THEN #temp_text1 := ' ';  END_IF;

